      Visibility <- "ST_HMI_Var_HMI_r64Axis_ChengXing_Position_real2"
   Line "线_346" at 68,549 size 180x6
      Visibility <- "ST_HMI_Var_HMI_r64Axis_ChengXing_Position_real2"
   Line "线_29" at 68,549 size 180x9
      Visibility <- "ST_HMI_Var_HMI_r64Axis_ChengXing_Position_real2"
   Line "线_31" at 68,549 size 166x68
      Visibility <- "ST_HMI_Var_HMI_r64Axis_ChengXing_Position_real2"
   Line "线_136#mig1_1" at 68,549 size 132x120
      Visibility <- "ST_HMI_Var_HMI_r64Axis_ChengXing_Position_real2"
   Line "线_38" at 68,443 size 144x106
      Visibility <- "ST_HMI_Var_HMI_r64Axis_ChengXing_Position_real2"
   Line "线_39" at 68,497 size 172x52
      Visibility <- "ST_HMI_Var_HMI_r64Axis_ChengXing_Position_real2"
   Line "线_11#mig1_1" at 68,441 size 143x108
      Visibility <- "ST_HMI_Var_HMI_r64Axis_ChengXing_Position_real2"
   Line "线_41" at 68,501 size 173x48
      Visibility <- "ST_HMI_Var_HMI_r64Axis_ChengXing_Position_real2"
   Line "线_43" at 68,549 size 129x122
      Visibility <- "ST_HMI_Var_HMI_r64Axis_ChengXing_Position_real2"
   Line "线_44" at 68,446 size 146x103
      Visibility <- "ST_HMI_Var_HMI_r64Axis_ChengXing_Position_real2"
   Line "线_115#mig1_1" at 68,549 size 179x13
      Visibility <- "ST_HMI_Var_HMI_r64Axis_ChengXing_Position_real2"
   Line "线_46" at 68,549 size 165x71
      Visibility <- "ST_HMI_Var_HMI_r64Axis_ChengXing_Position_real2"
   Line "线_47" at 68,549 size 179x15
      Visibility <- "ST_HMI_Var_HMI_r64Axis_ChengXing_Position_real2"
   Line "线_48" at 68,549 size 163x74
      Visibility <- "ST_HMI_Var_HMI_r64Axis_ChengXing_Position_real2"
   Line "线_49" at 68,549 size 127x124
      Visibility <- "ST_HMI_Var_HMI_r64Axis_ChengXing_Position_real2"
   Line "线_13#mig1_1" at 68,448 size 147x101
      Visibility <- "ST_HMI_Var_HMI_r64Axis_ChengXing_Position_real2"
   Line "线_59" at 68,503 size 174x46
      Visibility <- "ST_HMI_Var_HMI_r64Axis_ChengXing_Position_real2"
   Line "线_60" at 68,549 size 179x18
      Visibility <- "ST_HMI_Var_HMI_r64Axis_ChengXing_Position_real2"
   Line "线_61" at 68,549 size 162x77
      Visibility <- "ST_HMI_Var_HMI_r64Axis_ChengXing_Position_real2"
   Line "线_65" at 68,549 size 125x126
      Visibility <- "ST_HMI_Var_HMI_r64Axis_ChengXing_Position_real2"
   Line "线_124#mig1_1" at 68,451 size 149x98
      Visibility <- "ST_HMI_Var_HMI_r64Axis_ChengXing_Position_real2"
   Line "线_66" at 68,507 size 175x42
      Visibility <- "ST_HMI_Var_HMI_r64Axis_ChengXing_Position_real2"
   Line "线_67" at 68,549 size 179x21
      Visibility <- "ST_HMI_Var_HMI_r64Axis_ChengXing_Position_real2"
   Line "线_69" at 68,549 size 161x80
      Visibility <- "ST_HMI_Var_HMI_r64Axis_ChengXing_Position_real2"
   Line "线_70" at 68,549 size 122x129
      Visibility <- "ST_HMI_Var_HMI_r64Axis_ChengXing_Position_real2"
   Line "线_71" at 68,454 size 151x95
      Visibility <- "ST_HMI_Var_HMI_r64Axis_ChengXing_Position_real2"
   Line "线_72" at 68,510 size 175x39
      Visibility <- "ST_HMI_Var_HMI_r64Axis_ChengXing_Position_real2"
   Line "线_73" at 68,549 size 178x24
      Visibility <- "ST_HMI_Var_HMI_r64Axis_ChengXing_Position_real2"
   Line "线_74" at 68,549 size 159x82
      Visibility <- "ST_HMI_Var_HMI_r64Axis_ChengXing_Position_real2"
   Line "线_76" at 68,549 size 120x131
      Visibility <- "ST_HMI_Var_HMI_r64Axis_ChengXing_Position_real2"
   Line "线_77" at 68,456 size 153x93
      Visibility <- "ST_HMI_Var_HMI_r64Axis_ChengXing_Position_real2"
   Line "线_78" at 68,513 size 176x36
      Visibility <- "ST_HMI_Var_HMI_r64Axis_ChengXing_Position_real2"
   Line "线_79" at 68,549 size 178x27
      Visibility <- "ST_HMI_Var_HMI_r64Axis_ChengXing_Position_real2"
   Line "线_82" at 68,549 size 157x85
      Visibility <- "ST_HMI_Var_HMI_r64Axis_ChengXing_Position_real2"
   Line "线_84" at 68,549 size 118x133
      Visibility <- "ST_HMI_Var_HMI_r64Axis_ChengXing_Position_real2"
   Line "线_86" at 68,459 size 154x90
      Visibility <- "ST_HMI_Var_HMI_r64Axis_ChengXing_Position_real2"
   Line "线_87" at 68,516 size 177x33
      Visibility <- "ST_HMI_Var_HMI_r64Axis_ChengXing_Position_real2"
   Line "线_88" at 68,549 size 177x31
      Visibility <- "ST_HMI_Var_HMI_r64Axis_ChengXing_Position_real2"
   Line "线_90" at 68,549 size 156x88
      Visibility <- "ST_HMI_Var_HMI_r64Axis_ChengXing_Position_real2"
   Line "线_92" at 68,549 size 116x135
      Visibility <- "ST_HMI_Var_HMI_r64Axis_ChengXing_Position_real2"
   Line "线_93" at 68,462 size 156x87
      Visibility <- "ST_HMI_Var_HMI_r64Axis_ChengXing_Position_real2"
   Line "线_125#mig1_1" at 68,518 size 177x31
      Visibility <- "ST_HMI_Var_HMI_r64Axis_ChengXing_Position_real2"
   Line "线_98" at 68,549 size 177x33
      Visibility <- "ST_HMI_Var_HMI_r64Axis_ChengXing_Position_real2"
   Line "线_99" at 68,549 size 154x90
      Visibility <- "ST_HMI_Var_HMI_r64Axis_ChengXing_Position_real2"
   Line "线_109" at 68,549 size 113x137
      Visibility <- "ST_HMI_Var_HMI_r64Axis_ChengXing_Position_real2"
   Line "线_117" at 68,464 size 157x85
      Visibility <- "ST_HMI_Var_HMI_r64Axis_ChengXing_Position_real2"
   Line "线_119" at 68,521 size 178x28
      Visibility <- "ST_HMI_Var_HMI_r64Axis_ChengXing_Position_real2"
   Line "线_132" at 68,549 size 176x37
      Visibility <- "ST_HMI_Var_HMI_r64Axis_ChengXing_Position_real2"
   Line "线_135" at 68,549 size 153x93
      Visibility <- "ST_HMI_Var_HMI_r64Axis_ChengXing_Position_real2"
   Line "线_138" at 68,549 size 111x139
      Visibility <- "ST_HMI_Var_HMI_r64Axis_ChengXing_Position_real2"
   Line "线_347" at 68,466 size 159x83
      Visibility <- "ST_HMI_Var_HMI_r64Axis_ChengXing_Position_real2"
   Line "线_348" at 68,524 size 179x25
      Visibility <- "ST_HMI_Var_HMI_r64Axis_ChengXing_Position_real2"
   Line "线_349" at 68,549 size 175x39
      Visibility <- "ST_HMI_Var_HMI_r64Axis_ChengXing_Position_real2"
   Line "线_350" at 68,549 size 151x96
      Visibility <- "ST_HMI_Var_HMI_r64Axis_ChengXing_Position_real2"
   Line "线_351" at 68,549 size 108x141
      Visibility <- "ST_HMI_Var_HMI_r64Axis_ChengXing_Position_real2"
   Line "线_352" at 68,469 size 161x80
      Visibility <- "ST_HMI_Var_HMI_r64Axis_ChengXing_Position_real2"
   Line "线_130#mig1_1" at 68,527 size 179x22
      Visibility <- "ST_HMI_Var_HMI_r64Axis_ChengXing_Position_real2"
   Line "线_353" at 68,549 size 106x143
      Visibility <- "ST_HMI_Var_HMI_r64Axis_ChengXing_Position_real2"
   Line "线_97#mig1_1" at 68,471 size 162x78
      Visibility <- "ST_HMI_Var_HMI_r64Axis_ChengXing_Position_real2"
   Line "线_129#mig1_1" at 68,530 size 179x19
      Visibility <- "ST_HMI_Var_HMI_r64Axis_ChengXing_Position_real2"
   Line "线_354" at 68,549 size 175x43
      Visibility <- "ST_HMI_Var_HMI_r64Axis_ChengXing_Position_real2"
   Line "线_355" at 68,549 size 149x98
      Visibility <- "ST_HMI_Var_HMI_r64Axis_ChengXing_Position_real2"
   Line "线_356" at 68,549 size 103x144
      Visibility <- "ST_HMI_Var_HMI_r64Axis_ChengXing_Position_real2"
   Line "线_357" at 68,474 size 163x75
      Visibility <- "ST_HMI_Var_HMI_r64Axis_ChengXing_Position_real2"
   Line "线_128#mig1_1" at 68,534 size 179x15
      Visibility <- "ST_HMI_Var_HMI_r64Axis_ChengXing_Position_real2"
   Line "线_358" at 68,549 size 174x46
      Visibility <- "ST_HMI_Var_HMI_r64Axis_ChengXing_Position_real2"
   Line "线_359" at 68,549 size 147x101
      Visibility <- "ST_HMI_Var_HMI_r64Axis_ChengXing_Position_real2"
   Line "线_360" at 68,477 size 165x72
      Visibility <- "ST_HMI_Var_HMI_r64Axis_ChengXing_Position_real2"
   Line "线_131#mig1_1" at 68,536 size 179x13
      Visibility <- "ST_HMI_Var_HMI_r64Axis_ChengXing_Position_real2"
   Line "线_361" at 68,549 size 173x49
      Visibility <- "ST_HMI_Var_HMI_r64Axis_ChengXing_Position_real2"
   Line "线_362" at 68,549 size 146x104
      Visibility <- "ST_HMI_Var_HMI_r64Axis_ChengXing_Position_real2"
   Line "线_114#mig1_1" at 68,480 size 166x69
      Visibility <- "ST_HMI_Var_HMI_r64Axis_ChengXing_Position_real2"
   Line "线_363" at 68,540 size 180x9
      Visibility <- "ST_HMI_Var_HMI_r64Axis_ChengXing_Position_real2"
   Line "线_364" at 68,549 size 172x52
      Visibility <- "ST_HMI_Var_HMI_r64Axis_ChengXing_Position_real2"
   Line "线_365" at 68,549 size 144x106
      Visibility <- "ST_HMI_Var_HMI_r64Axis_ChengXing_Position_real2"
   Line "线_120#mig1_1" at 68,483 size 167x66
      Visibility <- "ST_HMI_Var_HMI_r64Axis_ChengXing_Position_real2"
   Line "线_366" at 68,543 size 180x6
      Visibility <- "ST_HMI_Var_HMI_r64Axis_ChengXing_Position_real2"
   Line "线_367" at 68,549 size 171x55
      Visibility <- "ST_HMI_Var_HMI_r64Axis_ChengXing_Position_real2"
   Line "线_368" at 68,549 size 142x109
      Visibility <- "ST_HMI_Var_HMI_r64Axis_ChengXing_Position_real2"
   Line "线_369" at 68,486 size 168x63
      Visibility <- "ST_HMI_Var_HMI_r64Axis_ChengXing_Position_real2"
   Line "线_150#mig1_1" at 68,546 size 180x3
      Visibility <- "ST_HMI_Var_HMI_r64Axis_ChengXing_Position_real2"
   Line "线_370" at 68,549 size 170x58
      Visibility <- "ST_HMI_Var_HMI_r64Axis_ChengXing_Position_real2"
   Line "线_371" at 68,549 size 140x111
      Visibility <- "ST_HMI_Var_HMI_r64Axis_ChengXing_Position_real2"
   Line "线_372" at 68,489 size 169x60
      Visibility <- "ST_HMI_Var_HMI_r64Axis_ChengXing_Position_real2"
   Line "线_147#mig1_1" at 68,549 size 180x0
      Visibility <- "ST_HMI_Var_HMI_r64Axis_ChengXing_Position_real2"
   Line "线_373" at 68,549 size 169x61
      Visibility <- "ST_HMI_Var_HMI_r64Axis_ChengXing_Position_real2"
   Line "线_374" at 68,549 size 138x114
      Visibility <- "ST_HMI_Var_HMI_r64Axis_ChengXing_Position_real2"
   Line "线_375" at 68,491 size 170x58
      Visibility <- "ST_HMI_Var_HMI_r64Axis_ChengXing_Position_real2"
   Line "线_376" at 68,549 size 180x3
      Visibility <- "ST_HMI_Var_HMI_r64Axis_ChengXing_Position_real2"
   Line "线_377" at 68,549 size 168x63
      Visibility <- "ST_HMI_Var_HMI_r64Axis_ChengXing_Position_real2"
   Line "线_378" at 68,549 size 167x67
      Visibility <- "ST_HMI_Var_HMI_r64Axis_ChengXing_Position_real2"
   Line "线_379" at 68,549 size 136x116
      Visibility <- "ST_HMI_Var_HMI_r64Axis_ChengXing_Position_real2"
   Line "线_380" at 68,549 size 134x118
      Visibility <- "ST_HMI_Var_HMI_r64Axis_ChengXing_Position_real2"
   Line "线_381" at 68,495 size 171x54
      Visibility <- "ST_HMI_Var_HMI_r64Axis_ChengXing_Position_real2"
   Line "线_382" at 68,549 size 180x6
      Visibility <- "ST_HMI_Var_HMI_r64Axis_ChengXing_Position_real2"
   ScreenModuleView "面板_1(2)_1" at 275,295 size 222x318; ScreenModuleType ""
      DirectMovement <- "ST_HMI_Var_HMI_r64Axis_ZouChe_Position_real2"
   Group "Group" at 136,477 size 84x252
   Polygon "多边形_8" at 152,627 size 24x54
      Visibility <- "VBS_hengsi_status0"
   Polygon "多边形_7" at 148,617 size 36x64
      Visibility <- "VBS_hengsi_status0"
   Polygon "多边形_10" at 146,607 size 42x74
      Visibility <- "VBS_hengsi_status0"
   Polygon "多边形_11#mig1" at 146,599 size 46x82
      Visibility <- "VBS_hengsi_status0"
   Polygon "多边形_12" at 144,591 size 52x90
      Visibility <- "VBS_hengsi_status0"
   Polygon "多边形_18" at 144,581 size 52x100
      Visibility <- "VBS_hengsi_status1"
   Polygon "多边形_17" at 144,573 size 56x108
      Visibility <- "VBS_hengsi_status1"
   Polygon "多边形_16" at 146,561 size 58x120
      Visibility <- "VBS_hengsi_status1"
   Polygon "多边形_15" at 146,549 size 62x134
      Visibility <- "VBS_hengsi_status1"
   Polygon "多边形_14" at 146,539 size 64x144
      Visibility <- "VBS_hengsi_status1"
   Polygon "多边形_19" at 144,529 size 68x154
      Visibility <- "VBS_hengsi_status1"
   Polygon "多边形_20" at 146,515 size 70x168
      Visibility <- "VBS_hengsi_status1"
   Polygon "多边形_21" at 144,509 size 74x174
      Visibility <- "VBS_hengsi_status1"
   Polygon "多边形_22" at 144,503 size 76x180
      Visibility <- "VBS_hengsi_status1"
   Group "Group_11" at 2,441 size 263x129
   Group "Group_6" at 0,523 size 86x54
   Group "Group_9" at 2,441 size 263x129
   Group "Group_10" at 2,441 size 263x129
   Line "线_10" at 32,520 size 233x8
      Visibility <- "ST_HMI_Var_HMI_r64Axis_1_ZhangLi_Position_JuanRao_real2"
   Line "线_12" at 32,528 size 233x0
      Visibility <- "ST_HMI_Var_HMI_r64Axis_1_ZhangLi_Position_JuanRao_real2"
   Line "线_17" at 32,524 size 233x4
      Visibility <- "ST_HMI_Var_HMI_r64Axis_1_ZhangLi_Position_JuanRao_real2"
   Line "线_18" at 32,528 size 233x4
      Visibility <- "ST_HMI_Var_HMI_r64Axis_1_ZhangLi_Position_JuanRao_real2"
   Line "线_19" at 32,528 size 233x8
      Visibility <- "ST_HMI_Var_HMI_r64Axis_1_ZhangLi_Position_JuanRao_real2"
   Line "线_20" at 32,528 size 233x12
      Visibility <- "ST_HMI_Var_HMI_r64Axis_1_ZhangLi_Position_JuanRao_real2"
   Line "线_116" at 32,528 size 232x16
      Visibility <- "ST_HMI_Var_HMI_r64Axis_1_ZhangLi_Position_JuanRao_real2"
   Line "线_118" at 32,528 size 232x21
      Visibility <- "ST_HMI_Var_HMI_r64Axis_1_ZhangLi_Position_JuanRao_real2"
   Line "线_121" at 32,528 size 232x25
      Visibility <- "ST_HMI_Var_HMI_r64Axis_1_ZhangLi_Position_JuanRao_real2"
   Line "线_126" at 32,528 size 231x29
      Visibility <- "ST_HMI_Var_HMI_r64Axis_1_ZhangLi_Position_JuanRao_real2"
   Line "线_127" at 32,528 size 231x33
      Visibility <- "ST_HMI_Var_HMI_r64Axis_1_ZhangLi_Position_JuanRao_real2"
   Line "线_128" at 32,441 size 216x87
      Visibility <- "ST_HMI_Var_HMI_r64Axis_1_ZhangLi_Position_JuanRao_real2"
   Line "线_129" at 32,445 size 218x83
      Visibility <- "ST_HMI_Var_HMI_r64Axis_1_ZhangLi_Position_JuanRao_real2"
   Line "线_130" at 32,448 size 219x80
      Visibility <- "ST_HMI_Var_HMI_r64Axis_1_ZhangLi_Position_JuanRao_real2"
   Line "线_131" at 32,452 size 220x76
      Visibility <- "ST_HMI_Var_HMI_r64Axis_1_ZhangLi_Position_JuanRao_real2"
   Line "线_133" at 32,456 size 222x72
      Visibility <- "ST_HMI_Var_HMI_r64Axis_1_ZhangLi_Position_JuanRao_real2"
   Line "线_134" at 32,460 size 223x68
      Visibility <- "ST_HMI_Var_HMI_r64Axis_1_ZhangLi_Position_JuanRao_real2"
   Line "线_136" at 32,464 size 224x64
      Visibility <- "ST_HMI_Var_HMI_r64Axis_1_ZhangLi_Position_JuanRao_real2"
   Line "线_137" at 32,468 size 225x60
      Visibility <- "ST_HMI_Var_HMI_r64Axis_1_ZhangLi_Position_JuanRao_real2"
   Line "线_139" at 32,472 size 226x56
      Visibility <- "ST_HMI_Var_HMI_r64Axis_1_ZhangLi_Position_JuanRao_real2"
   Line "线_140" at 32,476 size 227x52
      Visibility <- "ST_HMI_Var_HMI_r64Axis_1_ZhangLi_Position_JuanRao_real2"
   Line "线_141" at 32,480 size 228x48
      Visibility <- "ST_HMI_Var_HMI_r64Axis_1_ZhangLi_Position_JuanRao_real2"
   Line "线_142" at 32,484 size 229x44
      Visibility <- "ST_HMI_Var_HMI_r64Axis_1_ZhangLi_Position_JuanRao_real2"
   Line "线_143" at 32,488 size 230x40
      Visibility <- "ST_HMI_Var_HMI_r64Axis_1_ZhangLi_Position_JuanRao_real2"
   Line "线_144" at 32,492 size 230x36
      Visibility <- "ST_HMI_Var_HMI_r64Axis_1_ZhangLi_Position_JuanRao_real2"
   Line "线_145" at 32,496 size 231x32
      Visibility <- "ST_HMI_Var_HMI_r64Axis_1_ZhangLi_Position_JuanRao_real2"
   Line "线_146" at 32,500 size 231x28
      Visibility <- "ST_HMI_Var_HMI_r64Axis_1_ZhangLi_Position_JuanRao_real2"
   Line "线_147" at 32,504 size 232x24
      Visibility <- "ST_HMI_Var_HMI_r64Axis_1_ZhangLi_Position_JuanRao_real2"
   Line "线_148" at 32,507 size 232x21
      Visibility <- "ST_HMI_Var_HMI_r64Axis_1_ZhangLi_Position_JuanRao_real2"
   Line "线_149" at 32,512 size 232x16
      Visibility <- "ST_HMI_Var_HMI_r64Axis_1_ZhangLi_Position_JuanRao_real2"
   Line "线_150" at 32,516 size 233x12
      Visibility <- "ST_HMI_Var_HMI_r64Axis_1_ZhangLi_Position_JuanRao_real2"
   Line "线_151" at 32,520 size 233x8
      Visibility <- "ST_HMI_Var_HMI_r64Axis_1_ZhangLi_Position_JuanRao_real2"
   Line "线_152" at 32,528 size 233x0
      Visibility <- "ST_HMI_Var_HMI_r64Axis_1_ZhangLi_Position_JuanRao_real2"
   Line "线_153" at 32,524 size 233x4
      Visibility <- "ST_HMI_Var_HMI_r64Axis_1_ZhangLi_Position_JuanRao_real2"
   Line "线_154" at 32,528 size 233x4
      Visibility <- "ST_HMI_Var_HMI_r64Axis_1_ZhangLi_Position_JuanRao_real2"
   Line "线_155" at 32,528 size 233x8
      Visibility <- "ST_HMI_Var_HMI_r64Axis_1_ZhangLi_Position_JuanRao_real2"
   Line "线_156" at 32,528 size 233x12
      Visibility <- "ST_HMI_Var_HMI_r64Axis_1_ZhangLi_Position_JuanRao_real2"
   Line "线_158" at 32,528 size 232x16
      Visibility <- "ST_HMI_Var_HMI_r64Axis_1_ZhangLi_Position_JuanRao_real2"
   Line "线_160" at 32,528 size 232x21
      Visibility <- "ST_HMI_Var_HMI_r64Axis_1_ZhangLi_Position_JuanRao_real2"
   Line "线_161" at 32,528 size 232x25
      Visibility <- "ST_HMI_Var_HMI_r64Axis_1_ZhangLi_Position_JuanRao_real2"
   Line "线_162" at 32,528 size 231x29
      Visibility <- "ST_HMI_Var_HMI_r64Axis_1_ZhangLi_Position_JuanRao_real2"
   Line "线_163" at 32,528 size 231x33
      Visibility <- "ST_HMI_Var_HMI_r64Axis_1_ZhangLi_Position_JuanRao_real2"
   Line "线_164" at 32,441 size 216x87
      Visibility <- "ST_HMI_Var_HMI_r64Axis_1_ZhangLi_Position_JuanRao_real2"
   Line "线_165" at 32,445 size 218x83
      Visibility <- "ST_HMI_Var_HMI_r64Axis_1_ZhangLi_Position_JuanRao_real2"
   Line "线_166" at 32,448 size 219x80
      Visibility <- "ST_HMI_Var_HMI_r64Axis_1_ZhangLi_Position_JuanRao_real2"
   Line "线_167" at 32,452 size 220x76
      Visibility <- "ST_HMI_Var_HMI_r64Axis_1_ZhangLi_Position_JuanRao_real2"
   Line "线_168" at 32,456 size 222x72
      Visibility <- "ST_HMI_Var_HMI_r64Axis_1_ZhangLi_Position_JuanRao_real2"
   Line "线_169" at 32,460 size 223x68
      Visibility <- "ST_HMI_Var_HMI_r64Axis_1_ZhangLi_Position_JuanRao_real2"
   Line "线_170" at 32,464 size 224x64
      Visibility <- "ST_HMI_Var_HMI_r64Axis_1_ZhangLi_Position_JuanRao_real2"
   Line "线_171" at 32,468 size 225x60
      Visibility <- "ST_HMI_Var_HMI_r64Axis_1_ZhangLi_Position_JuanRao_real2"
   Line "线_172" at 32,472 size 226x56
      Visibility <- "ST_HMI_Var_HMI_r64Axis_1_ZhangLi_Position_JuanRao_real2"
   Line "线_173" at 32,476 size 227x52
      Visibility <- "ST_HMI_Var_HMI_r64Axis_1_ZhangLi_Position_JuanRao_real2"
   Line "线_174" at 32,480 size 228x48
      Visibility <- "ST_HMI_Var_HMI_r64Axis_1_ZhangLi_Position_JuanRao_real2"
   Line "线_175" at 32,484 size 229x44
      Visibility <- "ST_HMI_Var_HMI_r64Axis_1_ZhangLi_Position_JuanRao_real2"
   Line "线_176" at 32,488 size 230x40
      Visibility <- "ST_HMI_Var_HMI_r64Axis_1_ZhangLi_Position_JuanRao_real2"
   Line "线_177" at 32,492 size 230x36
      Visibility <- "ST_HMI_Var_HMI_r64Axis_1_ZhangLi_Position_JuanRao_real2"
   Line "线_178" at 32,496 size 231x32
      Visibility <- "ST_HMI_Var_HMI_r64Axis_1_ZhangLi_Position_JuanRao_real2"
   Line "线_179" at 32,500 size 231x28
      Visibility <- "ST_HMI_Var_HMI_r64Axis_1_ZhangLi_Position_JuanRao_real2"
   Line "线_180" at 32,504 size 232x24
      Visibility <- "ST_HMI_Var_HMI_r64Axis_1_ZhangLi_Position_JuanRao_real2"
   Line "线_181" at 32,507 size 232x21
      Visibility <- "ST_HMI_Var_HMI_r64Axis_1_ZhangLi_Position_JuanRao_real2"
   Line "线_182" at 32,512 size 232x16
      Visibility <- "ST_HMI_Var_HMI_r64Axis_1_ZhangLi_Position_JuanRao_real2"
   Line "线_183" at 32,516 size 233x12
      Visibility <- "ST_HMI_Var_HMI_r64Axis_1_ZhangLi_Position_JuanRao_real2"
   Group "Group_7" at 301,546 size 184x46
      DirectMovement <- "ST_HMI_Var_HMI_r64Axis_ZouChe_Position_real2"
   Group "Group_12" at 1030,614 size 136x46
   TextField "文本域_1" at 435,546 size 50x42; Text 'mm'
   IOField "IO Field_51" at 301,546 size 134x46; FormatPattern 9999.9
      ProcessValue <- "ST_HMI_Var_HMI_r64Axis_ZouChe_Position_real"
   TextField "文本域_2" at 1129,614 size 37x42; Text 'mm'
   IOField "IO Field_1" at 1030,614 size 99x46; FormatPattern 9999.9
      ProcessValue <- "ST_HMI_Var_HMI_r64_ZouChe_ZhanJu_Max_Effect"

screen "设置画面" 1280x733, template "模板_2"
   on GenerateScreen: function_b456aad1(1, N); SetTag("变量_100", 3)
   TextField "Text Field_25" at 26,537 size 151x33; Text '总牵伸: / 総ドラフト: / 전체 드라프트:'
   TextField "Text Field_26" at 26,608 size 151x34; Text '送条牵伸: / 篠送出しドラフト: / 담프롤러 드라프트:'
   TextField "Text Field_28" at 321,608 size 180x34; Text '第一牵伸(3段): / 第一ドラフト（3段）: / 제1드라프트(3단):'
   TextField "Text Field_37" at 304,679 size 197x34; Text '集中牵伸区(3段): / 集中ドラフトゾーン（3段）: / 집중 드라프트 구역(3단):'
   TextField "Text Field_38" at 321,537 size 180x33; Text '第一牵伸区(3段): / 第一ドラフトゾーン（3段）: / 제1드라프트 구역(3단):'
   TextField "Text Field_39" at 626,537 size 47x33; Text 'mm'
   TextField "Text Field_42" at 626,676 size 33x34; Text 'mm'
   TextField "Text Field_27" at 8,679 size 169x34; Text '分散牵伸(2段): / 分散ドラフト（2段）: / 캐리지드라프트(2단):'
   SymbolicIOField "符号 IO 域_1" at 186,466 size 121x40; TextOn '1'; TextOff '0'; TextList "QainShen_Select"
      ProcessValue <- "ST_HMI_Var_HMI_i16_QianShen_Select"
   IOField "IO Field_14" at 186,533 size 121x40; FormatPattern 9.99
      ProcessValue <- "ST_HMI_Var_HMI_r64QianShen_All"
   IOField "IO Field_15" at 186,605 size 121x40; FormatPattern 9.999
      ProcessValue <- "ST_HMI_Var_HMI_r64QianShen_WuNian"
   IOField "IO Field_17" at 502,605 size 121x40; FormatPattern 9.99
      ProcessValue <- "ST_HMI_Var_HMI_r64QianShen_First"
   IOField "IO Field_20" at 502,677 size 121x40; FormatPattern 99
      ProcessValue <- "ST_HMI_Var_HMI_r64QianShen_finalArea"
   IOField "IO Field_21" at 502,533 size 121x40; FormatPattern 999
      ProcessValue <- "ST_HMI_Var_HMI_r64QianShen_FirstArea"
   IOField "IO Field_16" at 186,677 size 121x40; FormatPattern 9.99
      ProcessValue <- "ST_HMI_Var_HMI_r64QianShen_FenSan"
   TextField "Text Field_19" at 695,20 size 137x38; Text '捻缩捻度: ジャッキング．イン 開始撚数: 작킹모션'
   TextField "Text Field_20" at 695,85 size 137x38; Text '捻缩距离: ジャッキング．イン 距離: 연축거리:'
   TextField "Text Field_21" at 695,150 size 137x38; Text '捻缩时间: ジャッキング．イン 時間: 연축시간:'
   TextField "Text Field_22" at 695,215 size 137x38; Text '捻缩速度: ジャッキング．イン 速度: 연축속도:'
   TextField "Text Field_31" at 695,285 size 130x32; Text '卷绕长度: / 巻取長: / 와인딩 길이:'
   TextField "Text Field_32" at 970,24 size 63x32; Text 'T/M'
   TextField "Text Field_33" at 970,89 size 63x32; Text 'mm'
   TextField "Text Field_35" at 970,219 size 63x32; Text 'mm/s'
   TextField "Text Field_36" at 970,285 size 63x32; Text 'mm'
   IOField "IO Field_11" at 839,150 size 121x40; FormatPattern 99.9
      ProcessValue <- "ST_HMI_Var_HMI_r64Time_NianSuo"
   IOField "IO Field_12" at 839,215 size 121x40; FormatPattern 99.9
      ProcessValue <- "ST_HMI_Var_HMI_r64Velocity_NianSuo"
      Appearance <- "ST_HMI_Var_HMI_boAlarm_NianSuo_SuDuOver"
   IOField "IO Field_19" at 839,281 size 121x40; FormatPattern 9999
      ProcessValue <- "ST_HMI_Var_HMI_r64Length_JuanRao"
   TextField "Text Field_41" at 724,597 size 132x31; Text '纱穗个数: / コップ本数: / 코프갯수:'
   TextField "Text Field_41#mig1" at 724,671 size 132x31; Text '单纱张力: / 単糸張力: / 단사 장력:'
   IOField "IO Field_75" at 867,594 size 121x40; FormatPattern 9999
      ProcessValue <- "ST_HMI_Var_HMI_r64_ShuLiang_ShaSui"
   IOField "IO Field_76" at 867,667 size 121x40; FormatPattern 999.9
      ProcessValue <- "ST_HMI_Var_HMI_r64_LuoSha_Force_DanSha_ZhangLi_FangKai"
   Button "OBJECT_106" at 1074,2 size 205x42; TextOff '手动 / EXIT / 手動 / 수동'; TextList "mode_enabled_1"
      ProcessValue <- "ST_Main_Var_g_i16_Mode_Enabled"
      Appearance <- "ST_Main_Var_g_i16_Mode_Enabled"
   Button "OBJECT_111" at 1074,45 size 205x42; TextOff '手动 / EXIT / 手動 / 수동'; TextList "automatic_status_1"
      Visibility <- "ST_Main_Var_g_bo_Mode_Enabled_Automatic"
      ProcessValue <- "ST_Main_Var_g_i16_Automatic_Status"
      Appearance <- "ST_Main_Var_g_i16_Automatic_Status"
   TextField "文本域_5" at 61,442 size 880x170; Text '锭子不转报警！请至报警画面解除报警，然后点击“退 出紧急停止”，点击“启动”开机，或者按正常步骤断电 重启，然后开机 捻度报警！设置捻度为 ， 实际捻度为 ， 已自动停止，请检查设置画面参数，重新设置总捻度， 检查设置其他参数，使画面上的参数没有红色闪烁，然 后按“启动”，若继续出现此报警，请从生头重新开始 스핀들이 돌아가지 않아 경보알림! 경보알림화면으로 이동하여 경보 해제후 "종료 비상 정지"를 클릭후 "시 작"을 클릭하여 가동하거나 정상적인 순서대로 단전 및 재부팅후 가동한다.'
      Visibility <- "ST_HMI_Var_HMI_i16_Dingzi_50102AlarmStatus"
   TextField "Text Field_5" at 615,155 size 60x32; Text 'r/min'
   IOField "IO Field_2" at 488,151 size 121x40; FormatPattern 99999
      ProcessValue <- "ST_HMI_Var_HMI_r64NianSu_Max"
      Appearance <- "ST_HMI_Var_HMI_boAlarm_NianDu_Time"
   TextField "Text Field_13" at 328,155 size 70x32; Text 'mm/s'
   TextField "Text Field_4" at 15,157 size 176x31; Text '出车速度: / 出機速度: / 외진속도:'
   TextField "Text Field_3" at 15,85 size 176x38; Text '牵伸捻度匹配值: ドラフト撚数マッチン グ値: 트위스트 연도 매칭값:'
   Button "OBJECT_107" at 416,216 size 230x40; TextOn '追捻启用 / 追撚使用 / 헤드 트위스트 사용'; TextOff '追捻启用 / EXIT / 追撚使用 / 헤드 트위스트 사용'
      Appearance <- "ST_HMI_Var_HMI_boNianDu_3"
   Button "OBJECT_1" at 416,280 size 230x40; TextOn '追捻停用 / 追撚停止 / 헤드 트위스트 사용중지'; TextOff '追捻停用 / EXIT / 追撚停止 / 헤드 트위스트 사용중지'
      Appearance <- "ST_HMI_Var_HMI_boNianDu_3"
   TextField "Text Field_9" at 15,216 size 176x38; Text '追捻开始捻度: / 追撚開始撚数: / 2단 요리 시작:'
   TextField "Text Field_10" at 328,220 size 70x32; Text 'T/M'
   TextField "Text Field_11" at 328,285 size 70x32; Text 'r/min'
   TextField "Text Field_16" at 81,384 size 101x30; Text '进车速度: / 入機速度: / 내진속도:'
   IOField "IO Field_22" at 186,379 size 121x40; FormatPattern 9999
      on OnFinishInput: SetBit("ST_Calculation_Var_HMI_bo_Calculation_0_Start"); SetTag("ST_Calculation_Var_g_i16_Calculation_0_3_Select_Status", 1)
      ProcessValue <- "ST_HMI_Var_HMI_r64Velocity_JinChe"
   TextField "Text Field_17" at 319,383 size 70x32; Text 'mm/s'
   TextField "Text Field_18" at 368,384 size 124x30; Text '展距: / 展開距離: / 스트레치 거리:'
   IOField "IO Field_23" at 492,379 size 121x40; FormatPattern 9999
      on OnFinishInput: SetBit("ST_Calculation_Var_HMI_bo_Calculation_0_Start"); SetTag("ST_Calculation_Var_g_i16_Calculation_0_3_Select_Status", 1)
      ProcessValue <- "ST_HMI_Var_HMI_r64Position_ChuChe"
   TextField "Text Field_23" at 617,383 size 32x32; Text 'mm'
   TextField "Text Field_24" at 15,282 size 176x38; Text '追捻锭子速度: 追撚スピンドル回転数: 헤드 트위스트 스핀들 속도:'
   TextField "Text Field_8" at 724,526 size 132x31; Text '纱穗直径: / コップ直径: / 코프 직경:'
   TextField "Text Field_29" at 385,25 size 101x30; Text '支数: / 番手: / 번수:'
   IOField "IO Field_24" at 867,521 size 121x40; FormatPattern 99.9
      on OnFinishInput: SetBit("ST_Calculation_Var_HMI_bo_Calculation_0_Start"); SetTag("ST_Calculation_Var_g_i16_Calculation_0_3_Select_Status", 1)
      ProcessValue <- "ST_HMI_Var_HMI_r64Diameter_ShaSui_Max"
   TextField "Text Field_14" at 993,525 size 70x32; Text 'mm'
   TextField "Text Field_2" at 15,25 size 176x31; Text '总捻度: / 総撚数: / 전체 연도:'
   TextField "Text Field_6" at 328,25 size 70x32; Text 'T/M'
   IOField "IO Field_13" at 488,85 size 121x40; FormatPattern 99.9
      ProcessValue <- "ST_HMI_Var_HMI_r64Time_JiaNian"
      Appearance <- "ST_HMI_Var_HMI_boAlarm_NianDu_Time"
   Button "HmiScreenItemData_3" at 1106,375 size 145x54; TextOn '纱穗参数设定 / 코핑 매개변수 설정'; TextOff '纱穗参数设定 / 코핑 매개변수 설정'
   Button "HmiScreenItemData_2" at 1106,275 size 145x54; TextOn '车况设定'; TextOff '车况设定'
   Button "HmiScreenItemData_1" at 1106,176 size 145x54; TextOn '向后 / 後向き / 뒤로'; TextOff '向后 / 後向き / 뒤로'
      on Release: ActivateScreen("自动画面", 0); function_f23ef4c9()
   TextField "Text Field_48" at 615,89 size 52x32; Text 's'
   TextField "Text Field_7" at 615,23 size 60x32; Text 'Nm'
   Button "按钮_5" at 894,361 size 147x69; TextOn '我要保存配方 / レシピを保存する / 레시피 저장'; TextOff '我要保存配方 / レシピを保存する / 레시피 저장'
      on Click: ActivateScreen("配方保存画面", 0)
   Button "按钮_2" at 714,361 size 147x69; TextOn '我要选择配方 / レシピを選択する / 레시피 선택'; TextOff '我要选择配方 / レシピを選択する / 레시피 선택'
      on Click: ActivateScreen("配方选择画面", 0)
   IOField "IO Field_1" at 195,85 size 121x40; FormatPattern 999
      on OnFinishInput: SetBit("ST_Calculation_Var_HMI_bo_Calculation_0_Start"); SetTag("ST_Calculation_Var_g_i16_Calculation_0_3_Select_Status", 1)
      ProcessValue <- "ST_HMI_Var_HMI_r64NianDu_QianShen_Best"
   IOField "IO Field_7" at 195,151 size 121x40; FormatPattern 9999
      on OnFinishInput: SetBit("ST_Calculation_Var_HMI_bo_Calculation_0_Start"); SetTag("ST_Calculation_Var_g_i16_Calculation_0_3_Select_Status", 1)
      ProcessValue <- "ST_HMI_Var_HMI_r64Velocity_ChuChe"
   IOField "IO Field_4" at 195,216 size 121x40; FormatPattern 9999
      on OnFinishInput: SetBit("ST_Calculation_Var_HMI_bo_Calculation_0_Start"); SetTag("ST_Calculation_Var_g_i16_Calculation_0_3_Select_Status", 1)
      ProcessValue <- "ST_HMI_Var_HMI_r64NianDu_1"
   IOField "IO Field_5" at 195,282 size 121x40; FormatPattern 99999
      on OnFinishInput: SetBit("ST_Calculation_Var_HMI_bo_Calculation_0_Start"); SetTag("ST_Calculation_Var_g_i16_Calculation_0_3_Select_Status", 1)
      ProcessValue <- "ST_HMI_Var_HMI_r64NianSu_2"
   IOField "IO Field_18" at 488,20 size 121x40; FormatPattern 99.9
      ProcessValue <- "ST_HMI_Var_HMI_r64ZhiShu_ChengSha"
   IOField "IO Field_43" at 195,20 size 121x40; FormatPattern 9999
      on OnFinishInput: SetBit("ST_Calculation_Var_HMI_bo_Calculation_0_Start"); SetTag("ST_Calculation_Var_g_i16_Calculation_0_3_Select_Status", 1)
      ProcessValue <- "ST_HMI_Var_HMI_r64NianDu_all"
   IOField "IO Field_3" at 839,20 size 121x40; FormatPattern 9999
      ProcessValue <- "ST_HMI_Var_HMI_r64NianDu_NianSuo"
   IOField "IO Field_6" at 839,85 size 121x40; FormatPattern 999
      ProcessValue <- "ST_HMI_Var_HMI_r64Position_NianSuo"
      Appearance <- "ST_HMI_Var_HMI_boAlarm_NianSuo_PosNon"
   Button "HmiScreenItemData_4" at 1106,479 size 145x54; TextOn '高级设置 / エキスパート設定 / 고급 설정'; TextOff '高级设置 / エキスパート設定 / 고급 설정'
      on Release: ActivateScreen("常用调试画面", 0)
   TextField "Text Field_34" at 970,154 size 63x33; Text 's'
   TextField "Text Field_1" at 392,85 size 94x38; Text '加捻时间: / 撚掛時間: / 연사시간:'
   TextField "Text Field_12" at 392,151 size 94x38; Text '锭子速度: スピンドル 回転数: 스핀들속도:'
   Button "HmiScreenItemData_5" at 1106,334 size 145x54; TextOn '高级设置 / エキスパート設定 / 고급 설정'; TextOff '监控画面 / エキスパート設定 / 고급 설정'
      on Release: ActivateScreen("监控画面", 0)
   Button "按钮_12" at 838,20 size 121x40; TextOff 'Text'
      on Click: ActivateScreen("参数修改画面", 0)
   Button "按钮_13" at 838,85 size 121x40; TextOff 'Text'
      on Click: ActivateScreen("参数修改画面", 0)
   Button "按钮_11" at 487,20 size 121x40; TextOff 'Text'
      on Click: ActivateScreen("参数修改画面", 0)
   Button "按钮_10" at 192,281 size 121x40; TextOff 'Text'
      on Click: ActivateScreen("参数修改画面", 0)
   Button "按钮_9" at 192,215 size 121x40; TextOff 'Text'
      on Click: ActivateScreen("参数修改画面", 0)
   Button "按钮_8" at 192,150 size 121x40; TextOff 'Text'
      on Click: ActivateScreen("参数修改画面", 0)
   Button "按钮_7" at 192,85 size 121x40; TextOff 'Text'
      on Click: ActivateScreen("参数修改画面", 0)
   Button "按钮_1" at 192,20 size 121x40; TextOff 'Text'
      on Click: ActivateScreen("参数修改画面", 0)
   Button "按钮_16" at 751,544 size 137x44; TextOff '知道了 / OK'
      on Click: SetTag("ST_HMI_Var_HMI_i16_Dingzi_50102AlarmStatus", 0); ResetBit("ST_HMI_Var_HMI_bo_XiangLing")
      Visibility <- "ST_HMI_Var_HMI_i16_Dingzi_50102AlarmStatus"
   Circle "圆_3" at 791,455 size 60x60
      Visibility <- "ST_HMI_Var_HMI_i16_Dingzi_50102AlarmStatus"
      Appearance <- "ST_HMI_Var_HMI_bo_XiangLing"
   TextField "文本域_11" at 12,427 size 880x170; Text '捻度报警！设置捻度为 ， 实际捻度为 ， 已自动停止，请检查设置画面参数，重新设置总捻度， 检查设置其他参数，使画面上的参数没有红色闪烁，然 后按“启动”，若继续出现此报警，请从生头重新开始 트위스트 경보 알림!설정 트위스트는 이고,실제 트위스트는 이며, 이미 자동정지, 설정화면 매개변수를 확인하고, 전체 트위스트를 다 시 설정하고, 기타 매개변수를 확인설정하여 화면의 매개변수에 빨간색이 깜빡이지 않도록 해야 한다. 그다음 "작동"을 누른다. 만약 이 경보가 연속 반복적으로 나타나면 스레딩부터 다시 시작한다.'
      Visibility <- "ST_HMI_Var_HMI_i16_NianduAlarmStatus"
   IOField "IO Field_8" at 388,428 size 86x32; FormatPattern 9999
      on OnFinishInput: SetBit("ST_Calculation_Var_HMI_bo_Calculation_0_Start"); SetTag("ST_Calculation_Var_g_i16_Calculation_0_3_Select_Status", 1)
      Visibility <- "ST_HMI_Var_HMI_i16_NianduAlarmStatus"
      ProcessValue <- "ST_HMI_Var_HMI_r64NianDu_all"
   IOField "IO Field_9" at 699,428 size 86x32; FormatPattern 9999
      Visibility <- "ST_HMI_Var_HMI_i16_NianduAlarmStatus"
      ProcessValue <- "ST_HMI_Var_HMI_r64Niandu_all_Current"
   Button "按钮_6" at 745,537 size 137x44; TextOff '知道了 / OK'
      on Click: SetTag("ST_HMI_Var_HMI_i16_NianduAlarmStatus", 0); SetBit("ST_Calculation_Var_HMI_bo_Calculation_0_Start"); ResetBit("ST_HMI_Var_HMI_bo_XiangLing")
      Visibility <- "ST_HMI_Var_HMI_i16_NianduAlarmStatus"
   Circle "圆_2" at 785,448 size 60x60
      Visibility <- "ST_HMI_Var_HMI_i16_NianduAlarmStatus"
      Appearance <- "ST_HMI_Var_HMI_bo_XiangLing"

